// TIA Portal project "OPCUA_S71x00" (V16)

(* hardware
DEVICE "S71500/ET200MP station_2"  S7-1500 station
   slot 0: "Rail_0"  Rack  6ES7 590-1***0-0AA0
   slot 1: "1511f"  CPU 1511F-1 PN  6ES7 511-1FK02-0AB0  V2.8
      slot 3: "CPU display_1"  6ES7591-1AA00-0AA0
      slot 32768: "PROFINET interface_1"  X1
         slot 32769: "Port_1"  X1 P1
         slot 32770: "Port_2"  X1 P2
      slot 34817: "Virtual CP interface port_1"  Virtual CP interface port  Virtual CP interface port
DEVICE "S7-1200 station_2"  S7-1200 Station
   slot 0: "Rack_0"  S7-1200 Rack  Rack  V1.0
   slot 1: "1212fc"  CPU 1212FC DC/DC/DC  6ES7 212-1AF40-0XB0  V4.4
DEVICE "S7-1200 station_1"  S7-1200 Station
   slot 0: "Rack_0"  S7-1200 Rack  Rack  V1.0
   slot 1: "1214c"  CPU 1214C DC/DC/DC  6ES7 214-1AG40-0XB0  V4.4
*)

// ===== PLC "1511f"  CPU 1511F-1 PN =====

VAR_GLOBAL   // PLC tag table "Default tag table"
   "Tag_1" AT %MW0 : Int;
   "Tag_2" AT %MW2 : Int;
   "tag_bool" AT %M4.0 : Bool;
   "tab_byte" AT %MB6 : Byte;
   "tag_int" AT %MW7 : Int;
   "Tag_3" AT %MW4 : Int;
   "Tag_4" AT %MW6 : Int;
END_VAR

DATA_BLOCK "db_opcua"   // DB2
{ S7_Optimized_Access := 'TRUE' }
VERSION : 0.1
   VAR
      zm_array : Array[0..2] of Byte;
      zm_bool : Bool;
      zm_byte : Byte;
      zm_char : Char;
      zm_datetime_date_and_time : Date_And_Time;
      zm_datetime_dtl : DTL;
      zm_dword : DWord;
      zm_int : Int;
      zm_datetime_ldt : LDT;
      zm_real : Real;
      zm_string : String;
      zm_struct : Struct
         zm_struct_bool : Bool;
         zm_struct_byte : Byte;
      END_STRUCT;
   END_VAR
BEGIN
END_DATA_BLOCK

ORGANIZATION_BLOCK "Main"   // OB1, LAD, ProgramCycle
TITLE = "Main Program Sweep (Cycle)"
{ S7_Optimized_Access := 'TRUE' }
VERSION : 0.1
   VAR_INPUT
      Initial_Call : Bool;   // Initial call of this OB
      Remanence : Bool;   // =True, if remanent data are available
   END_VAR
BEGIN

REGION Network 1
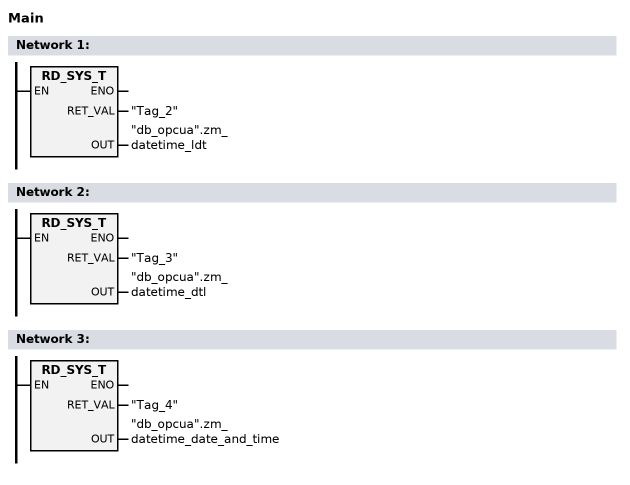
   "Tag_2" := RD_SYS_T(OUT => "db_opcua".zm_datetime_ldt);
END_REGION

REGION Network 2
   "Tag_3" := RD_SYS_T(OUT => "db_opcua".zm_datetime_dtl);
END_REGION

REGION Network 3
   "Tag_4" := RD_SYS_T(OUT => "db_opcua".zm_datetime_date_and_time);
END_REGION
END_ORGANIZATION_BLOCK

// ===== PLC "1212fc"  CPU 1212FC DC/DC/DC =====

VAR_GLOBAL   // PLC tag table "Default tag table"
   "Tag_1" AT %MW0 : Int;
   "set_ctu" AT %M2.0 : Bool;
   "reset_ctu" AT %M2.1 : Bool;
END_VAR

DATA_BLOCK "db_opcua"   // DB1
{ S7_Optimized_Access := 'TRUE' }
VERSION : 0.1
   VAR
      zm_array : Array[0..2] of Byte;
      zm_bool : Bool;
      zm_byte : Byte;
      zm_char : Char;
      zm_datetime_dtl : DTL;
      zm_dword : DWord;
      zm_int : Int;
      zm_real : Real;
      zm_string : String;
      zm_struct : Struct
         zm_struct_bool : Bool;
         zm_struct_byte : Byte;
      END_STRUCT;
   END_VAR
BEGIN
END_DATA_BLOCK

// folder: System blocks/Program resources

DATA_BLOCK "IEC_Counter_0_DB"   // DB2
{ S7_Optimized_Access := 'TRUE' }
AUTHOR : Simatic
FAMILY : IEC
NAME : CNTR
VERSION : 1.0
// stored: InstanceOfName IEC_COUNTER
"IEC_COUNTER"
BEGIN
END_DATA_BLOCK

// folder: (top level)

ORGANIZATION_BLOCK "Main"   // OB1, LAD, ProgramCycle
TITLE = "Main Program Sweep (Cycle)"
{ S7_Optimized_Access := 'TRUE' }
VERSION : 0.1
   VAR_INPUT
      Initial_Call : Bool;   // Initial call of this OB
      Remanence : Bool;   // =True, if remanent data are available
   END_VAR
BEGIN

REGION Network 1
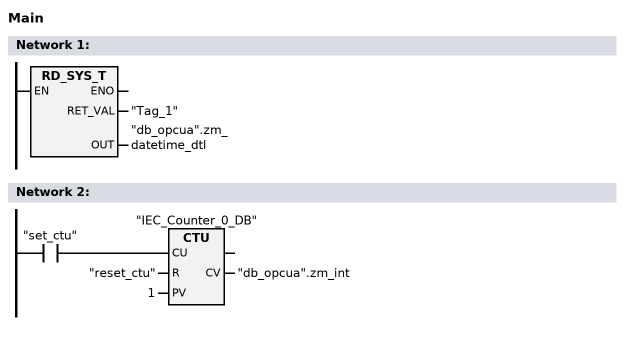
   "Tag_1" := RD_SYS_T(OUT => "db_opcua".zm_datetime_dtl);
END_REGION

REGION Network 2
   "IEC_Counter_0_DB".CTU(CU := "set_ctu", R := "reset_ctu", PV := 1, CV => "db_opcua".zm_int);
END_REGION
END_ORGANIZATION_BLOCK

// ===== PLC "1214c"  CPU 1214C DC/DC/DC =====

VAR_GLOBAL   // PLC tag table "Default tag table"
   "Tag_1" AT %MW0 : Int;
   "set_ctu" AT %M2.0 : Bool;
   "reset_ctu" AT %M2.1 : Bool;
END_VAR

DATA_BLOCK "db_opcua"   // DB1
{ S7_Optimized_Access := 'TRUE' }
VERSION : 0.1
   VAR
      zm_array : Array[0..2] of Byte;
      zm_bool : Bool;
      zm_byte : Byte;
      zm_char : Char;
      zm_datetime_dtl : DTL;
      zm_dword : DWord;
      zm_int : Int;
      zm_real : Real;
      zm_string : String;
      zm_struct : Struct
         zm_struct_bool : Bool;
         zm_struct_byte : Byte;
      END_STRUCT;
   END_VAR
BEGIN
END_DATA_BLOCK

// folder: System blocks/Program resources

DATA_BLOCK "IEC_Counter_0_DB"   // DB2
{ S7_Optimized_Access := 'TRUE' }
AUTHOR : Simatic
FAMILY : IEC
NAME : CNTR
VERSION : 1.0
// stored: InstanceOfName IEC_COUNTER
"IEC_COUNTER"
BEGIN
END_DATA_BLOCK

// folder: (top level)

ORGANIZATION_BLOCK "Main"   // OB1, LAD, ProgramCycle
TITLE = "Main Program Sweep (Cycle)"
{ S7_Optimized_Access := 'TRUE' }
VERSION : 0.1
   VAR_INPUT
      Initial_Call : Bool;   // Initial call of this OB
      Remanence : Bool;   // =True, if remanent data are available
   END_VAR
BEGIN

REGION Network 1
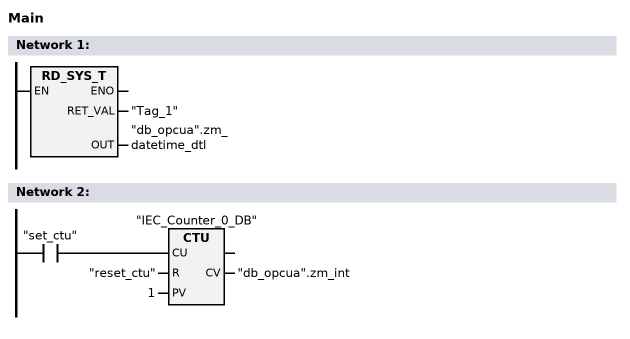
   "Tag_1" := RD_SYS_T(OUT => "db_opcua".zm_datetime_dtl);
END_REGION

REGION Network 2
   "IEC_Counter_0_DB".CTU(CU := "set_ctu", R := "reset_ctu", PV := 1, CV => "db_opcua".zm_int);
END_REGION
END_ORGANIZATION_BLOCK